
screen "AI" 800x480, template "Main"
   Button "Button_1" at 7,5 size 96x32; TextOff 'Мешалки'; Authorization "Admin"
      on Release: ActivateScreen("Mix", 0); SetTag("settings", 1)
      Appearance <- "settings"
   Button "Button_2" at 7,52 size 96x32; TextOff 'Дозаторы'; Authorization "Admin"
      on Release: ActivateScreen("Dos", 0); SetTag("settings", 2)
      Appearance <- "settings"
   Button "Button_3" at 7,99 size 96x32; TextOff 'Клапана'; Authorization "Admin"
      on Release: ActivateScreen("Valve", 0); SetTag("settings", 3)
      Appearance <- "settings"
   Button "Button_4" at 7,146 size 96x32; TextOff 'AI'; Authorization "Admin"
      on Release: ActivateScreen("AI", 0); SetTag("settings", 4)
      Appearance <- "settings"
   Button "Button_5" at 7,193 size 96x32; TextOff 'DI'; Authorization "Admin"
      on Release: ActivateScreen("DI", 0); SetTag("settings", 5)
      Appearance <- "settings"
   Button "Button_6" at 7,240 size 96x32; TextOff 'DO'; Authorization "Admin"
      on Release: ActivateScreen("DO", 0); SetTag("settings", 6)
      Appearance <- "settings"
   TextField "Text field_2" at 210,15 size 67x22; Text 'Датчик:'
   TextField "Text field_4" at 282,15 size 99x22; Text 'Расходомер'
   TextField "Text field_7" at 390,18 size 43x22; Text 'вход'
   TextField "Text field_8" at 390,43 size 56x22; Text 'выход'
   IOField "I/O field_1" at 456,19 size 92x26; FormatPattern s999999999.999
      ProcessValue <- "AIx_DB_FlowMeter_Converter_Min_In"
   IOField "I/O field_2" at 456,41 size 92x26; FormatPattern s999999999.999
      ProcessValue <- "AIx_DB_FlowMeter_Converter_Min_Out"
   IOField "I/O field_3" at 555,18 size 92x26; FormatPattern s999999999.999
      ProcessValue <- "AIx_DB_FlowMeter_Converter_Max_In"
   IOField "I/O field_4" at 555,40 size 92x26; FormatPattern s999999999.999
      ProcessValue <- "AIx_DB_FlowMeter_Converter_Max_Out"
   TextField "Text field_9" at 389,68 size 101x22; Text 'Фильтрация'
   TextField "Text field_10" at 390,96 size 36x22; Text 'RTD'
   Button "Button_7" at 489,71 size 20x20; TextOff 'Text'; PictureList "ok"
      on Click: InvertBit("AIx_DB_FlowMeter_Use_Filter")
      ProcessValue <- "AIx_DB_FlowMeter_Use_Filter"
   Button "Button_8" at 489,96 size 20x20; TextOff 'Text'; PictureList "ok"
      on Click: InvertBit("AIx_DB_FlowMeter_Use_RTD")
      ProcessValue <- "AIx_DB_FlowMeter_Use_RTD"
   IOField "I/O field_5" at 516,68 size 65x25; FormatPattern 999
      ProcessValue <- "AIx_DB_FlowMeter_Filter_SP"
   IOField "I/O field_6" at 516,93 size 65x25; FormatPattern 999
      ProcessValue <- "AIx_DB_FlowMeter_RTD_c"
   TextField "Text field_11" at 210,36 size 79x22; Text 'Поправка'
   IOField "I/O field_7" at 293,36 size 78x23; FormatPattern s999.9
      ProcessValue <- "AIx_DB_FlowMeter_Calibration"
   Button "Button_9" at 396,176 size 248x28; TextOff 'Use'
      on Click: InvertBit("AIx_DB_FlowMeter_CMD_Start_A")
      Appearance <- "AIx_DB_FlowMeter_CMD_Start_A"
   Button "Button_10" at 213,66 size 68x28; TextOff 'Hand'
      on Click: InvertBit("AIx_DB_FlowMeter_CMD_Hand")
      Appearance <- "AIx_DB_FlowMeter_CMD_Hand"
   IOField "I/O field_8" at 293,66 size 78x28; FormatPattern s9999.9
      ProcessValue <- "AIx_DB_FlowMeter_Result"
   TextField "Text field_12" at 436,123 size 27x22; Text 'NC'
   TextField "Text field_13" at 437,143 size 25x22; Text 'SC'
   TextField "Text field_14" at 210,125 size 27x22; Text 'HH'
   TextField "Text field_15" at 216,145 size 16x22; Text 'H'
   TextField "Text field_16" at 217,165 size 14x22; Text 'L'
   TextField "Text field_17" at 212,186 size 23x22; Text 'LL'
   IOField "I/O field_11" at 472,123 size 58x21; FormatPattern s99999
      ProcessValue <- "AIx_DB_FlowMeter_SP_NC"
   IOField "I/O field_12" at 472,143 size 58x21; FormatPattern s99999
      ProcessValue <- "AIx_DB_FlowMeter_SP_SC"
   IOField "I/O field_13" at 246,125 size 58x21; FormatPattern 99999
      ProcessValue <- "AIx_DB_FlowMeter_SP_HH"
   IOField "I/O field_14" at 246,145 size 58x21; FormatPattern 99999
      ProcessValue <- "AIx_DB_FlowMeter_SP_H"
   IOField "I/O field_15" at 246,165 size 58x21; FormatPattern s99999
      ProcessValue <- "AIx_DB_FlowMeter_SP_L"
   IOField "I/O field_16" at 246,185 size 58x21; FormatPattern s99999
      ProcessValue <- "AIx_DB_FlowMeter_SP_LL"
   IOField "I/O field_17" at 546,123 size 58x21; FormatPattern 999
      ProcessValue <- "AIx_DB_FlowMeter_Timers_NC_SP"
   IOField "I/O field_18" at 546,143 size 58x21; FormatPattern 999
      ProcessValue <- "AIx_DB_FlowMeter_Timers_SC_SP"
   IOField "I/O field_19" at 320,125 size 58x21; FormatPattern 999
      ProcessValue <- "AIx_DB_FlowMeter_Timers_HH_SP"
   IOField "I/O field_20" at 320,145 size 58x21; FormatPattern 999
      ProcessValue <- "AIx_DB_FlowMeter_Timers_H_SP"
   IOField "I/O field_21" at 320,165 size 58x21; FormatPattern 999
      ProcessValue <- "AIx_DB_FlowMeter_Timers_L_SP"
   IOField "I/O field_22" at 320,185 size 58x21; FormatPattern 999
      ProcessValue <- "AIx_DB_FlowMeter_Timers_LL_SP"
   IOField "I/O field_23" at 582,93 size 65x25; FormatPattern s99999
      ProcessValue <- "AIx_DB_FlowMeter_Signal"
   TextField "Text field_18" at 210,97 size 68x22; Text 'Уставка'
   TextField "Text field_19" at 299,97 size 79x22; Text 'Время (с)'
   TextField "Text field_1" at 214,248 size 67x22; Text 'Датчик:'
   TextField "Text field_3" at 286,248 size 69x22; Text 'Уровень'
   TextField "Text field_5" at 394,251 size 43x22; Text 'вход'
   TextField "Text field_6" at 394,276 size 56x22; Text 'выход'
   IOField "I/O field_9" at 460,252 size 92x26; FormatPattern s999999999.999
      ProcessValue <- "AIx_DB_Level_Converter_Min_In"
   IOField "I/O field_10" at 460,274 size 92x26; FormatPattern s999999999.999
      ProcessValue <- "AIx_DB_Level_Converter_Min_Out"
   IOField "I/O field_24" at 559,251 size 92x26; FormatPattern s999999999.999
      ProcessValue <- "AIx_DB_Level_Converter_Max_In"
   IOField "I/O field_25" at 559,273 size 92x26; FormatPattern s999999999.999
      ProcessValue <- "AIx_DB_Level_Converter_Max_Out"
   TextField "Text field_20" at 393,301 size 101x22; Text 'Фильтрация'
   TextField "Text field_21" at 394,329 size 36x22; Text 'RTD'
   Button "Button_11" at 493,304 size 20x20; TextOff 'Text'; PictureList "ok"
      on Click: InvertBit("AIx_DB_Level_Use_Filter")
      ProcessValue <- "AIx_DB_Level_Use_Filter"
   Button "Button_12" at 493,329 size 20x20; TextOff 'Text'; PictureList "ok"
      on Click: InvertBit("AIx_DB_Level_Use_RTD")
      ProcessValue <- "AIx_DB_Level_Use_RTD"
   IOField "I/O field_26" at 520,301 size 65x25; FormatPattern 999
      ProcessValue <- "AIx_DB_Level_Filter_SP"
   IOField "I/O field_27" at 520,326 size 65x25; FormatPattern 999
      ProcessValue <- "AIx_DB_Level_RTD_c"
   TextField "Text field_22" at 214,269 size 79x22; Text 'Поправка'
   IOField "I/O field_28" at 297,269 size 78x23; FormatPattern s999.9
      ProcessValue <- "AIx_DB_Level_Calibration"
   Button "Button_13" at 400,409 size 248x28; TextOff 'Use'
      on Click: InvertBit("AIx_DB_Level_CMD_Start_A")
      Appearance <- "AIx_DB_Level_CMD_Start_A"
   Button "Button_14" at 217,299 size 68x28; TextOff 'Hand'
      on Click: InvertBit("AIx_DB_Level_CMD_Hand")
      Appearance <- "AIx_DB_Level_CMD_Hand"
   IOField "I/O field_29" at 297,299 size 78x28; FormatPattern s9999.9
      ProcessValue <- "AIx_DB_Level_Result"
   TextField "Text field_23" at 440,356 size 27x22; Text 'NC'
   TextField "Text field_24" at 441,376 size 25x22; Text 'SC'
   TextField "Text field_25" at 214,358 size 27x22; Text 'HH'
   TextField "Text field_26" at 220,378 size 16x22; Text 'H'
   TextField "Text field_27" at 221,398 size 14x22; Text 'L'
   TextField "Text field_28" at 216,419 size 23x22; Text 'LL'
   IOField "I/O field_30" at 476,356 size 58x21; FormatPattern s99999
      ProcessValue <- "AIx_DB_Level_SP_NC"
   IOField "I/O field_31" at 476,376 size 58x21; FormatPattern s99999
      ProcessValue <- "AIx_DB_Level_SP_SC"
   IOField "I/O field_32" at 250,358 size 58x21; FormatPattern 99999
      ProcessValue <- "AIx_DB_Level_SP_HH"
   IOField "I/O field_33" at 250,378 size 58x21; FormatPattern 99999
      ProcessValue <- "AIx_DB_Level_SP_H"
   IOField "I/O field_34" at 250,398 size 58x21; FormatPattern s99999
      ProcessValue <- "AIx_DB_Level_SP_L"
   IOField "I/O field_35" at 250,418 size 58x21; FormatPattern s99999
      ProcessValue <- "AIx_DB_Level_SP_LL"
   IOField "I/O field_36" at 550,356 size 58x21; FormatPattern 999
      ProcessValue <- "AIx_DB_Level_Timers_NC_SP"
   IOField "I/O field_37" at 550,376 size 58x21; FormatPattern 999
      ProcessValue <- "AIx_DB_Level_Timers_SC_SP"
   IOField "I/O field_38" at 324,358 size 58x21; FormatPattern 999
      ProcessValue <- "AIx_DB_Level_Timers_HH_SP"
   IOField "I/O field_39" at 324,378 size 58x21; FormatPattern 999
      ProcessValue <- "AIx_DB_Level_Timers_H_SP"
   IOField "I/O field_40" at 324,398 size 58x21; FormatPattern 999
      ProcessValue <- "AIx_DB_Level_Timers_L_SP"
   IOField "I/O field_41" at 324,418 size 58x21; FormatPattern 999
      ProcessValue <- "AIx_DB_Level_Timers_LL_SP"
   IOField "I/O field_42" at 586,326 size 65x25; FormatPattern s99999
      ProcessValue <- "AIx_DB_Level_Signal"
   TextField "Text field_29" at 214,330 size 68x22; Text 'Уставка'
   TextField "Text field_30" at 303,330 size 79x22; Text 'Время (с)'

screen "DI" 800x480, template "Main"
   Button "Button_1" at 7,5 size 96x32; TextOff 'Мешалки'; Authorization "Admin"
      on Release: ActivateScreen("Mix", 0); SetTag("settings", 1)
      Appearance <- "settings"
   Button "Button_2" at 7,52 size 96x32; TextOff 'Дозаторы'; Authorization "Admin"
      on Release: ActivateScreen("Dos", 0); SetTag("settings", 2)
      Appearance <- "settings"
   Button "Button_3" at 7,99 size 96x32; TextOff 'Клапана'; Authorization "Admin"
      on Release: ActivateScreen("Valve", 0); SetTag("settings", 3)
      Appearance <- "settings"
   Button "Button_4" at 7,146 size 96x32; TextOff 'AI'; Authorization "Admin"
      on Release: ActivateScreen("AI", 0); SetTag("settings", 4)
      Appearance <- "settings"
   Button "Button_5" at 7,193 size 96x32; TextOff 'DI'; Authorization "Admin"
      on Release: ActivateScreen("DI", 0); SetTag("settings", 5)
      Appearance <- "settings"
   Button "Button_6" at 7,240 size 96x32; TextOff 'DO'; Authorization "Admin"
      on Release: ActivateScreen("DO", 0); SetTag("settings", 6)
      Appearance <- "settings"
   Group "Group" at 127,7 size 283x51; TextList "Hand"
   Group "Group_1" at 127,66 size 283x51; TextList "Hand"
   Group "Group_2" at 127,125 size 283x51; TextList "Hand"
   Group "Group_3" at 127,184 size 283x51; TextList "Hand"
   Group "Group_4" at 127,244 size 283x51; TextList "Hand"
   Group "Group_5" at 127,303 size 283x51; TextList "Hand"
   Group "Group_6" at 127,362 size 283x51; TextList "Hand"
   Group "Group_7" at 127,422 size 283x51; TextList "Hand"
   Group "Group_8" at 433,7 size 283x51; TextList "Hand"
   Group "Group_9" at 433,66 size 283x51; TextList "Hand"
   Group "Group_10" at 433,125 size 283x51; TextList "Hand"
   Group "Group_11" at 433,184 size 283x51; TextList "Hand"
   Group "Group_12" at 433,244 size 283x51; TextList "Hand"
   Group "Group_13" at 433,303 size 283x51; TextList "Hand"
   TextField "Text field_1" at 131,10 size 45x22; Text 'I 0.0'
   TextField "Text field_2" at 176,10 size 120x22; Text 'M1 Готовность'
   Circle "Circle_1" at 131,33 size 22x22
      Appearance <- "DIx_DB_M1_FB_Ready_Input"
   Circle "Circle_2" at 154,33 size 22x22
      Appearance <- "DIx_DB_M1_FB_Ready_Signal"
   Button "Button_7" at 298,11 size 59x44; TextOff 'Авто'; TextList "Hand"
      on Click: InvertBit("DIx_DB_M1_FB_Ready_Hand")
      Appearance <- "DIx_DB_M1_FB_Ready_Hand"
      ProcessValue <- "DIx_DB_M1_FB_Ready_Hand"
   Button "Button_8" at 240,33 size 49x22; TextOff 'Выкл'
      on Click: ResetBit("DIx_DB_M1_FB_Ready_Start_M")
   Button "Button_12" at 184,33 size 47x22; TextOff 'Вкл'
      on Click: SetBit("DIx_DB_M1_FB_Ready_Start_M")
      Appearance <- "DIx_DB_M1_FB_Ready_Start_M"
   IOField "I/O field_6" at 360,33 size 23x22; FormatPattern 99
      ProcessValue <- "DIx_DB_M1_FB_Ready_Filter_On_SP"
   IOField "I/O field_7" at 383,33 size 23x22; FormatPattern 99
      ProcessValue <- "DIx_DB_M1_FB_Ready_Filter_Off_SP"
   Button "Button_9" at 360,10 size 46x20; TextOff 'Inv'
      on Click: InvertBit("DIx_DB_M1_FB_Ready_Inverse")
      Appearance <- "DIx_DB_M1_FB_Ready_Inverse"
   TextField "Text field_3" at 131,69 size 45x22; Text 'I 0.1'
   TextField "Text field_4" at 176,69 size 87x22; Text 'M1 Работа'
   Circle "Circle_3" at 131,92 size 22x22
      Appearance <- "DIx_DB_M1_FB_Run_Input"
   Circle "Circle_4" at 154,92 size 22x22
      Appearance <- "DIx_DB_M1_FB_Run_Signal"
   Button "Button_10" at 298,70 size 59x44; TextOff 'Авто'; TextList "Hand"
      on Click: InvertBit("DIx_DB_M1_FB_Run_Hand")
      Appearance <- "DIx_DB_M1_FB_Run_Hand"
      ProcessValue <- "DIx_DB_M1_FB_Run_Hand"
   Button "Button_11" at 240,92 size 49x22; TextOff 'Выкл'
      on Click: ResetBit("DIx_DB_M1_FB_Run_Start_M")
   Button "Button_13" at 184,92 size 47x22; TextOff 'Вкл'
      on Click: SetBit("DIx_DB_M1_FB_Run_Start_M")
      Appearance <- "DIx_DB_M1_FB_Run_Start_M"
   IOField "I/O field_1" at 360,92 size 23x22; FormatPattern 99
      ProcessValue <- "DIx_DB_M1_FB_Run_Filter_On_SP"
   IOField "I/O field_2" at 383,92 size 23x22; FormatPattern 99
      ProcessValue <- "DIx_DB_M1_FB_Run_Filter_Off_SP"
   Button "Button_14" at 360,69 size 46x20; TextOff 'Inv'
      on Click: InvertBit("DIx_DB_M1_FB_Run_Inverse")
      Appearance <- "DIx_DB_M1_FB_Run_Inverse"
   TextField "Text field_5" at 131,128 size 45x22; Text 'I 0.2'
   TextField "Text field_6" at 176,128 size 120x22; Text 'M2 Готовность'
   Circle "Circle_5" at 131,151 size 22x22
      Appearance <- "DIx_DB_M2_FB_Ready_Input"
   Circle "Circle_6" at 154,151 size 22x22
      Appearance <- "DIx_DB_M2_FB_Ready_Signal"
   Button "Button_15" at 298,129 size 59x44; TextOff 'Авто'; TextList "Hand"
      on Click: InvertBit("DIx_DB_M2_FB_Ready_Hand")
      Appearance <- "DIx_DB_M2_FB_Ready_Hand"
      ProcessValue <- "DIx_DB_M2_FB_Ready_Hand"
   Button "Button_16" at 240,151 size 49x22; TextOff 'Выкл'
      on Click: ResetBit("DIx_DB_M2_FB_Ready_Start_M")
   Button "Button_17" at 184,151 size 47x22; TextOff 'Вкл'
      on Click: SetBit("DIx_DB_M2_FB_Ready_Start_M")
      Appearance <- "DIx_DB_M2_FB_Ready_Start_M"
   IOField "I/O field_3" at 360,151 size 23x22; FormatPattern 99
      ProcessValue <- "DIx_DB_M2_FB_Ready_Filter_On_SP"
   IOField "I/O field_4" at 383,151 size 23x22; FormatPattern 99
      ProcessValue <- "DIx_DB_M2_FB_Ready_Filter_Off_SP"
   Button "Button_18" at 360,128 size 46x20; TextOff 'Inv'
      on Click: InvertBit("DIx_DB_M2_FB_Ready_Inverse")
      Appearance <- "DIx_DB_M2_FB_Ready_Inverse"
   TextField "Text field_7" at 131,187 size 45x22; Text 'I 0.3'
   TextField "Text field_8" at 176,187 size 87x22; Text 'M2 Работа'
   Circle "Circle_7" at 131,210 size 22x22
      Appearance <- "DIx_DB_M2_FB_Run_Input"
   Circle "Circle_8" at 154,210 size 22x22
      Appearance <- "DIx_DB_M2_FB_Run_Signal"
   Button "Button_19" at 298,188 size 59x44; TextOff 'Авто'; TextList "Hand"
      on Click: InvertBit("DIx_DB_M2_FB_Run_Hand")
      Appearance <- "DIx_DB_M2_FB_Run_Hand"
      ProcessValue <- "DIx_DB_M2_FB_Run_Hand"
   Button "Button_20" at 240,210 size 49x22; TextOff 'Выкл'
      on Click: ResetBit("DIx_DB_M2_FB_Run_Start_M")
   Button "Button_21" at 184,210 size 47x22; TextOff 'Вкл'
      on Click: SetBit("DIx_DB_M2_FB_Run_Start_M")
      Appearance <- "DIx_DB_M2_FB_Run_Start_M"
   IOField "I/O field_5" at 360,210 size 23x22; FormatPattern 99
      ProcessValue <- "DIx_DB_M2_FB_Run_Filter_On_SP"
   IOField "I/O field_8" at 383,210 size 23x22; FormatPattern 99
      ProcessValue <- "DIx_DB_M2_FB_Run_Filter_Off_SP"
   Button "Button_22" at 360,187 size 46x20; TextOff 'Inv'
      on Click: InvertBit("DIx_DB_M2_FB_Run_Inverse")
      Appearance <- "DIx_DB_M2_FB_Run_Inverse"
   TextField "Text field_9" at 131,247 size 45x22; Text 'I 0.4'
   TextField "Text field_10" at 176,247 size 120x22; Text 'M3 Готовность'
   Circle "Circle_9" at 131,270 size 22x22
      Appearance <- "DIx_DB_M3_FB_Ready_Input"
   Circle "Circle_10" at 154,270 size 22x22
      Appearance <- "DIx_DB_M3_FB_Ready_Signal"
   Button "Button_23" at 298,248 size 59x44; TextOff 'Авто'; TextList "Hand"
      on Click: InvertBit("DIx_DB_M3_FB_Ready_Hand")
      Appearance <- "DIx_DB_M3_FB_Ready_Hand"
      ProcessValue <- "DIx_DB_M3_FB_Ready_Hand"
   Button "Button_24" at 240,270 size 49x22; TextOff 'Выкл'
      on Click: ResetBit("DIx_DB_M3_FB_Ready_Start_M")
   Button "Button_25" at 184,270 size 47x22; TextOff 'Вкл'
      on Click: SetBit("DIx_DB_M3_FB_Ready_Start_M")
      Appearance <- "DIx_DB_M3_FB_Ready_Start_M"
   IOField "I/O field_9" at 360,270 size 23x22; FormatPattern 99
      ProcessValue <- "DIx_DB_M3_FB_Ready_Filter_On_SP"
   IOField "I/O field_10" at 383,270 size 23x22; FormatPattern 99
      ProcessValue <- "DIx_DB_M3_FB_Ready_Filter_Off_SP"
   Button "Button_26" at 360,247 size 46x20; TextOff 'Inv'
      on Click: InvertBit("DIx_DB_M3_FB_Ready_Inverse")
      Appearance <- "DIx_DB_M3_FB_Ready_Inverse"
   TextField "Text field_11" at 131,306 size 45x22; Text 'I 0.5'
   TextField "Text field_12" at 176,306 size 87x22; Text 'M3 Работа'
   Circle "Circle_11" at 131,329 size 22x22
      Appearance <- "DIx_DB_M3_FB_Run_Input"
   Circle "Circle_12" at 154,329 size 22x22
      Appearance <- "DIx_DB_M3_FB_Run_Signal"
   Button "Button_27" at 298,307 size 59x44; TextOff 'Авто'; TextList "Hand"
      on Click: InvertBit("DIx_DB_M3_FB_Run_Hand")
      Appearance <- "DIx_DB_M3_FB_Run_Hand"
      ProcessValue <- "DIx_DB_M3_FB_Run_Hand"
   Button "Button_28" at 240,329 size 49x22; TextOff 'Выкл'
      on Click: ResetBit("DIx_DB_M3_FB_Run_Start_M")
   Button "Button_29" at 184,329 size 47x22; TextOff 'Вкл'
      on Click: SetBit("DIx_DB_M3_FB_Run_Start_M")
      Appearance <- "DIx_DB_M3_FB_Run_Start_M"
   IOField "I/O field_11" at 360,329 size 23x22; FormatPattern 99
      ProcessValue <- "DIx_DB_M3_FB_Run_Filter_On_SP"
   IOField "I/O field_12" at 383,329 size 23x22; FormatPattern 99
      ProcessValue <- "DIx_DB_M3_FB_Run_Filter_Off_SP"
   Button "Button_30" at 360,306 size 46x20; TextOff 'Inv'
      on Click: InvertBit("DIx_DB_M3_FB_Run_Inverse")
      Appearance <- "DIx_DB_M3_FB_Run_Inverse"
   TextField "Text field_13" at 131,365 size 45x22; Text 'I 0.6'
   TextField "Text field_14" at 176,365 size 120x22; Text 'Сух.доз.Готов.'
   Circle "Circle_13" at 131,388 size 22x22
      Appearance <- "DIx_DB_DD_FB_Ready_Input"
   Circle "Circle_14" at 154,388 size 22x22
      Appearance <- "DIx_DB_DD_FB_Ready_Signal"
   Button "Button_31" at 298,366 size 59x44; TextOff 'Авто'; TextList "Hand"
      on Click: InvertBit("DIx_DB_DD_FB_Ready_Hand")
      Appearance <- "DIx_DB_DD_FB_Ready_Hand"
      ProcessValue <- "DIx_DB_DD_FB_Ready_Hand"
   Button "Button_32" at 240,388 size 49x22; TextOff 'Выкл'
      on Click: ResetBit("DIx_DB_DD_FB_Ready_Start_M")
   Button "Button_33" at 184,388 size 47x22; TextOff 'Вкл'
      on Click: SetBit("DIx_DB_DD_FB_Ready_Start_M")
      Appearance <- "DIx_DB_DD_FB_Ready_Start_M"
   IOField "I/O field_13" at 360,388 size 23x22; FormatPattern 99
      ProcessValue <- "DIx_DB_DD_FB_Ready_Filter_On_SP"
   IOField "I/O field_14" at 383,388 size 23x22; FormatPattern 99
      ProcessValue <- "DIx_DB_DD_FB_Ready_Filter_Off_SP"
   Button "Button_34" at 360,365 size 46x20; TextOff 'Inv'
      on Click: InvertBit("DIx_DB_DD_FB_Ready_Inverse")
      Appearance <- "DIx_DB_DD_FB_Ready_Inverse"
   TextField "Text field_15" at 131,425 size 45x22; Text 'I 0.7'
   TextField "Text field_16" at 176,425 size 98x22; Text 'Доз. Работа'
   Circle "Circle_15" at 131,448 size 22x22
      Appearance <- "DIx_DB_Dos_FB_Run_Input"
   Circle "Circle_16" at 154,448 size 22x22
      Appearance <- "DIx_DB_Dos_FB_Run_Signal"
   Button "Button_35" at 298,426 size 59x44; TextOff 'Авто'; TextList "Hand"
      on Click: InvertBit("DIx_DB_Dos_FB_Run_Hand")
      ProcessValue <- "DIx_DB_Dos_FB_Run_Hand"
      Appearance <- "DIx_DB_Dos_FB_Run_Hand"
   Button "Button_36" at 240,448 size 49x22; TextOff 'Выкл'
      on Click: ResetBit("DIx_DB_Dos_FB_Run_Start_M")
   Button "Button_37" at 184,448 size 47x22; TextOff 'Вкл'
      on Click: SetBit("DIx_DB_Dos_FB_Run_Start_M")
      Appearance <- "DIx_DB_Dos_FB_Run_Start_M"
   IOField "I/O field_15" at 360,448 size 23x22; FormatPattern 99
      ProcessValue <- "DIx_DB_Dos_FB_Run_Filter_On_SP"
   IOField "I/O field_16" at 383,448 size 23x22; FormatPattern 99
      ProcessValue <- "DIx_DB_Dos_FB_Run_Filter_Off_SP"
   Button "Button_38" at 360,425 size 46x20; TextOff 'Inv'
      on Click: InvertBit("DIx_DB_Dos_FB_Run_Inverse")
      Appearance <- "DIx_DB_Dos_FB_Run_Inverse"
   TextField "Text field_17" at 437,10 size 45x22; Text 'I 1.0'
   TextField "Text field_18" at 482,10 size 95x22; Text 'Сух.доз.Ур.'
   Circle "Circle_17" at 437,33 size 22x22
      Appearance <- "DIx_DB_DD_LLS_Input"
   Circle "Circle_18" at 460,33 size 22x22
      Appearance <- "DIx_DB_DD_LLS_Signal"
   Button "Button_39" at 604,11 size 59x44; TextOff 'Авто'; TextList "Hand"
      on Click: InvertBit("DIx_DB_DD_LLS_Hand")
      Appearance <- "DIx_DB_DD_LLS_Hand"
      ProcessValue <- "DIx_DB_DD_LLS_Hand"
   Button "Button_40" at 546,33 size 49x22; TextOff 'Выкл'
      on Click: ResetBit("DIx_DB_DD_LLS_Start_M")
   Button "Button_41" at 490,33 size 47x22; TextOff 'Вкл'
      on Click: SetBit("DIx_DB_DD_LLS_Start_M")
      Appearance <- "DIx_DB_DD_LLS_Start_M"
   IOField "I/O field_17" at 666,33 size 23x22; FormatPattern 99
      ProcessValue <- "DIx_DB_DD_LLS_Filter_On_SP"
   IOField "I/O field_18" at 689,33 size 23x22; FormatPattern 99
      ProcessValue <- "DIx_DB_DD_LLS_Filter_Off_SP"
   Button "Button_42" at 666,10 size 46x20; TextOff 'Inv'
      on Click: InvertBit("DIx_DB_DD_LLS_Inverse")
      Appearance <- "DIx_DB_DD_LLS_Inverse"
   TextField "Text field_19" at 437,69 size 45x22; Text 'I 1.1'
   TextField "Text field_20" at 482,69 size 104x22; Text 'Вибро Готов.'
   Circle "Circle_19" at 437,92 size 22x22
      Appearance <- "DIx_DB_Vibro_FB_Ready_Input"
   Circle "Circle_20" at 460,92 size 22x22
      Appearance <- "DIx_DB_Vibro_FB_Ready_Signal"
   Button "Button_43" at 604,70 size 59x44; TextOff 'Авто'; TextList "Hand"
      on Click: InvertBit("DIx_DB_Vibro_FB_Ready_Hand")
      Appearance <- "DIx_DB_Vibro_FB_Ready_Hand"
      ProcessValue <- "DIx_DB_Vibro_FB_Ready_Hand"
   Button "Button_44" at 546,92 size 49x22; TextOff 'Выкл'
      on Click: ResetBit("DIx_DB_Vibro_FB_Ready_Start_M")
   Button "Button_45" at 490,92 size 47x22; TextOff 'Вкл'
      on Click: SetBit("DIx_DB_Vibro_FB_Ready_Start_M")
      Appearance <- "DIx_DB_Vibro_FB_Ready_Start_M"
   IOField "I/O field_19" at 666,92 size 23x22; FormatPattern 99
      ProcessValue <- "DIx_DB_Vibro_FB_Ready_Filter_On_SP"
   IOField "I/O field_20" at 689,92 size 23x22; FormatPattern 99
      ProcessValue <- "DIx_DB_Vibro_FB_Ready_Filter_Off_SP"
   Button "Button_46" at 666,69 size 46x20; TextOff 'Inv'
      on Click: InvertBit("DIx_DB_Vibro_FB_Ready_Inverse")
      Appearance <- "DIx_DB_Vibro_FB_Ready_Inverse"
   TextField "Text field_21" at 437,128 size 45x22; Text 'I 1.2'
   TextField "Text field_22" at 482,128 size 112x22; Text 'Пневмотранс.'
   Circle "Circle_21" at 437,151 size 22x22
      Appearance <- "DIx_DB_Transporter_Input"
   Circle "Circle_22" at 460,151 size 22x22
      Appearance <- "DIx_DB_Transporter_Signal"
   Button "Button_47" at 604,129 size 59x44; TextOff 'Авто'; TextList "Hand"
      on Click: InvertBit("DIx_DB_Transporter_Hand")
      Appearance <- "DIx_DB_Transporter_Hand"
      ProcessValue <- "DIx_DB_Transporter_Hand"
   Button "Button_48" at 546,151 size 49x22; TextOff 'Выкл'
      on Click: ResetBit("DIx_DB_Transporter_Start_M")
   Button "Button_49" at 490,151 size 47x22; TextOff 'Вкл'
      on Click: SetBit("DIx_DB_Transporter_Start_M")
      Appearance <- "DIx_DB_Transporter_Start_M"
   IOField "I/O field_21" at 666,151 size 23x22; FormatPattern 99
      ProcessValue <- "DIx_DB_Transporter_Filter_On_SP"
   IOField "I/O field_22" at 689,151 size 23x22; FormatPattern 99
      ProcessValue <- "DIx_DB_Transporter_Filter_Off_SP"
   Button "Button_50" at 666,128 size 46x20; TextOff 'Inv'
      on Click: InvertBit("DIx_DB_Transporter_Inverse")
      Appearance <- "DIx_DB_Transporter_Inverse"
   TextField "Text field_23" at 437,187 size 45x22; Text 'I 1.3'
   TextField "Text field_24" at 482,187 size 128x22; Text 'Жид.доз.Готов.'
   Circle "Circle_23" at 437,210 size 22x22
      Appearance <- "DIx_DB_DL_FB_Ready_Input"
   Circle "Circle_24" at 460,210 size 22x22
      Appearance <- "DIx_DB_DL_FB_Ready_Signal"
   Button "Button_51" at 604,188 size 59x44; TextOff 'Авто'; TextList "Hand"
      on Click: InvertBit("DIx_DB_DL_FB_Ready_Hand")
      Appearance <- "DIx_DB_DL_FB_Ready_Hand"
      ProcessValue <- "DIx_DB_DL_FB_Ready_Hand"
   Button "Button_52" at 546,210 size 49x22; TextOff 'Выкл'
      on Click: ResetBit("DIx_DB_DL_FB_Ready_Start_M")
   Button "Button_53" at 490,210 size 47x22; TextOff 'Вкл'
      on Click: SetBit("DIx_DB_DL_FB_Ready_Start_M")
      Appearance <- "DIx_DB_DL_FB_Ready_Start_M"
   IOField "I/O field_23" at 666,210 size 23x22; FormatPattern 99
      ProcessValue <- "DIx_DB_DL_FB_Ready_Filter_On_SP"
   IOField "I/O field_24" at 689,210 size 23x22; FormatPattern 99
      ProcessValue <- "DIx_DB_DL_FB_Ready_Filter_Off_SP"
   Button "Button_54" at 666,187 size 46x20; TextOff 'Inv'
      on Click: InvertBit("DIx_DB_DL_FB_Ready_Inverse")
      Appearance <- "DIx_DB_DL_FB_Ready_Inverse"
   TextField "Text field_25" at 437,247 size 45x22; Text 'I 1.4'
   TextField "Text field_26" at 482,247 size 61x22; Text 'Проток'
   Circle "Circle_25" at 437,270 size 22x22
      Appearance <- "DIx_DB_Dry_Run_Input"
   Circle "Circle_26" at 460,270 size 22x22
      Appearance <- "DIx_DB_Dry_Run_Signal"
   Button "Button_55" at 604,248 size 59x44; TextOff 'Авто'; TextList "Hand"
      on Click: InvertBit("DIx_DB_Dry_Run_Hand")
      Appearance <- "DIx_DB_Dry_Run_Hand"
      ProcessValue <- "DIx_DB_Dry_Run_Hand"
   Button "Button_56" at 546,270 size 49x22; TextOff 'Выкл'
      on Click: ResetBit("DIx_DB_Dry_Run_Start_M")
   Button "Button_57" at 490,270 size 47x22; TextOff 'Вкл'
      on Click: SetBit("DIx_DB_Dry_Run_Start_M")
      Appearance <- "DIx_DB_Dry_Run_Start_M"
   IOField "I/O field_25" at 666,270 size 23x22; FormatPattern 99
      ProcessValue <- "DIx_DB_Dry_Run_Filter_On_SP"
   IOField "I/O field_26" at 689,270 size 23x22; FormatPattern 99
      ProcessValue <- "DIx_DB_Dry_Run_Filter_Off_SP"
   Button "Button_58" at 666,247 size 46x20; TextOff 'Inv'
      on Click: InvertBit("DIx_DB_Dry_Run_Inverse")
      Appearance <- "DIx_DB_Dry_Run_Inverse"
   TextField "Text field_27" at 437,306 size 45x22; Text 'I 1.5'
   TextField "Text field_28" at 482,306 size 70x22; Text 'Останов'
   Circle "Circle_27" at 437,329 size 22x22
      Appearance <- "DIx_DB_AllBlock_Input"
   Circle "Circle_28" at 460,329 size 22x22
      Appearance <- "DIx_DB_AllBlock_Signal"
   Button "Button_59" at 604,307 size 59x44; TextOff 'Авто'; TextList "Hand"
      on Click: InvertBit("DIx_DB_AllBlock_Hand")
      Appearance <- "DIx_DB_AllBlock_Hand"
      ProcessValue <- "DIx_DB_AllBlock_Hand"
   Button "Button_60" at 546,329 size 49x22; TextOff 'Выкл'
      on Click: ResetBit("DIx_DB_AllBlock_Start_M")
   Button "Button_61" at 490,329 size 47x22; TextOff 'Вкл'
      on Click: SetBit("DIx_DB_AllBlock_Start_M")
      Appearance <- "DIx_DB_AllBlock_Start_M"
   IOField "I/O field_27" at 666,329 size 23x22; FormatPattern 99
      ProcessValue <- "DIx_DB_AllBlock_Filter_On_SP"
   IOField "I/O field_28" at 689,329 size 23x22; FormatPattern 99
      ProcessValue <- "DIx_DB_AllBlock_Filter_Off_SP"
   Button "Button_62" at 666,306 size 46x20; TextOff 'Inv'
      on Click: InvertBit("DIx_DB_AllBlock_Inverse")
      Appearance <- "DIx_DB_AllBlock_Inverse"

screen "DO" 800x480, template "Main"
   Button "Button_1" at 7,5 size 96x32; TextOff 'Мешалки'; Authorization "Admin"
      on Release: ActivateScreen("Mix", 0); SetTag("settings", 1)
      Appearance <- "settings"
   Button "Button_2" at 7,52 size 96x32; TextOff 'Дозаторы'; Authorization "Admin"
      on Release: ActivateScreen("Dos", 0); SetTag("settings", 2)
      Appearance <- "settings"
   Button "Button_3" at 7,99 size 96x32; TextOff 'Клапана'; Authorization "Admin"
      on Release: ActivateScreen("Valve", 0); SetTag("settings", 3)
      Appearance <- "settings"
   Button "Button_4" at 7,146 size 96x32; TextOff 'AI'; Authorization "Admin"
      on Release: ActivateScreen("AI", 0); SetTag("settings", 4)
      Appearance <- "settings"
   Button "Button_5" at 7,193 size 96x32; TextOff 'DI'; Authorization "Admin"
      on Release: ActivateScreen("DI", 0); SetTag("settings", 5)
      Appearance <- "settings"
   Button "Button_6" at 7,240 size 96x32; TextOff 'DO'; Authorization "Admin"
      on Release: ActivateScreen("DO", 0); SetTag("settings", 6)
      Appearance <- "settings"
   Group "Group" at 127,7 size 283x51; TextList "Hand"
   Group "Group_1" at 127,66 size 283x51; Text 'Q 0.0'; TextList "Hand"
   Group "Group_2" at 127,125 size 283x51; Text 'Q 0.0'; TextList "Hand"
   Group "Group_3" at 127,184 size 283x51; Text 'Q 0.0'; TextList "Hand"
   Group "Group_4" at 127,244 size 283x51; Text 'Q 0.0'; TextList "Hand"
   Group "Group_5" at 127,303 size 283x51; Text 'Q 0.0'; TextList "Hand"
   Group "Group_6" at 127,362 size 283x51; Text 'Q 0.0'; TextList "Hand"
   Group "Group_7" at 127,422 size 283x51; Text 'Q 0.0'; TextList "Hand"
   Group "Group_8" at 433,7 size 283x51; Text 'Q 0.0'; TextList "Hand"
   Group "Group_9" at 433,66 size 283x51; Text 'Q 0.0'; TextList "Hand"
   TextField "Text field_4" at 131,10 size 45x22; Text 'Q 0.0'
   TextField "Text field_5" at 176,10 size 69x22; Text 'M1 Пуск'
   Circle "Circle_3" at 131,33 size 22x22
      Appearance <- "DOx_DB_M1_CMD_Start_A"
   Circle "Circle_4" at 154,33 size 22x22
      Appearance <- "DOx_DB_M1_CMD_Q"
   Button "Button_13" at 298,11 size 59x44; TextOff 'Авто'; TextList "Hand"
      on Click: InvertBit("DOx_DB_M1_CMD_Hand")
      Appearance <- "DOx_DB_M1_CMD_Hand"
      ProcessValue <- "DOx_DB_M1_CMD_Hand"
   Button "Button_14" at 240,33 size 49x22; TextOff 'Выкл'
      on Click: ResetBit("DOx_DB_M1_CMD_Start_M")
   Button "Button_15" at 184,33 size 47x22; TextOff 'Вкл'
      on Click: SetBit("DOx_DB_M1_CMD_Start_M")
      Appearance <- "DOx_DB_M1_CMD_Start_M"
   Button "Button_16" at 360,10 size 46x20; TextOff 'Inv'
      on Click: InvertBit("DOx_DB_M1_CMD_Inverse")
      Appearance <- "DOx_DB_M1_CMD_Inverse"
   Button "Button_17" at 360,35 size 46x20; TextOff 'Sim'
      on Click: InvertBit("DOx_DB_M1_CMD_Simulation")
      Appearance <- "DOx_DB_M1_CMD_Simulation"
   TextField "Text field_1" at 131,69 size 45x22; Text 'Q 0.1'
   TextField "Text field_2" at 176,69 size 69x22; Text 'M2 Пуск'
   Circle "Circle_1" at 131,92 size 22x22
      Appearance <- "DOx_DB_M2_CMD_Start_A"
   Circle "Circle_2" at 154,92 size 22x22
      Appearance <- "DOx_DB_M2_CMD_Q"
   Button "Button_7" at 298,70 size 59x44; TextOff 'Авто'; TextList "Hand"
      on Click: InvertBit("DOx_DB_M2_CMD_Hand")
      Appearance <- "DOx_DB_M2_CMD_Hand"
      ProcessValue <- "DOx_DB_M2_CMD_Hand"
   Button "Button_8" at 240,92 size 49x22; TextOff 'Выкл'
      on Click: ResetBit("DOx_DB_M2_CMD_Start_M")
   Button "Button_9" at 184,92 size 47x22; TextOff 'Вкл'
      on Click: SetBit("DOx_DB_M2_CMD_Start_M")
      Appearance <- "DOx_DB_M2_CMD_Start_M"
   Button "Button_10" at 360,69 size 46x20; TextOff 'Inv'
      on Click: InvertBit("DOx_DB_M2_CMD_Inverse")
      Appearance <- "DOx_DB_M2_CMD_Inverse"
   Button "Button_11" at 360,94 size 46x20; TextOff 'Sim'
      on Click: InvertBit("DOx_DB_M2_CMD_Simulation")
      Appearance <- "DOx_DB_M2_CMD_Simulation"
   TextField "Text field_3" at 131,128 size 45x22; Text 'Q 0.2'
   TextField "Text field_6" at 176,128 size 69x22; Text 'M3 Пуск'
   Circle "Circle_5" at 131,151 size 22x22
      Appearance <- "DOx_DB_M3_CMD_Start_A"
   Circle "Circle_6" at 154,151 size 22x22
      Appearance <- "DOx_DB_M3_CMD_Q"
   Button "Button_12" at 298,129 size 59x44; TextOff 'Авто'; TextList "Hand"
      on Click: InvertBit("DOx_DB_M3_CMD_Hand")
      Appearance <- "DOx_DB_M3_CMD_Hand"
      ProcessValue <- "DOx_DB_M3_CMD_Hand"
   Button "Button_18" at 240,151 size 49x22; TextOff 'Выкл'
      on Click: ResetBit("DOx_DB_M3_CMD_Start_M")
   Button "Button_19" at 184,151 size 47x22; TextOff 'Вкл'
      on Click: SetBit("DOx_DB_M3_CMD_Start_M")
      Appearance <- "DOx_DB_M3_CMD_Start_M"
   Button "Button_20" at 360,128 size 46x20; TextOff 'Inv'
      on Click: InvertBit("DOx_DB_M3_CMD_Inverse")
      Appearance <- "DOx_DB_M3_CMD_Inverse"
   Button "Button_21" at 360,153 size 46x20; TextOff 'Sim'
      on Click: InvertBit("DOx_DB_M3_CMD_Simulation")
      Appearance <- "DOx_DB_M3_CMD_Simulation"
   TextField "Text field_7" at 131,187 size 45x22; Text 'Q 0.3'
   TextField "Text field_8" at 176,187 size 109x22; Text 'Сух.Доз.Пуск'
   Circle "Circle_7" at 131,210 size 22x22
      Appearance <- "DOx_DB_DD_CMD_Start_A"
   Circle "Circle_8" at 154,210 size 22x22
      Appearance <- "DOx_DB_DD_CMD_Q"
   Button "Button_22" at 298,188 size 59x44; TextOff 'Авто'; TextList "Hand"
      on Click: InvertBit("DOx_DB_DD_CMD_Hand")
      Appearance <- "DOx_DB_DD_CMD_Hand"
      ProcessValue <- "DOx_DB_DD_CMD_Hand"
   Button "Button_23" at 240,210 size 49x22; TextOff 'Выкл'
      on Click: ResetBit("DOx_DB_DD_CMD_Start_M")
   Button "Button_24" at 184,210 size 47x22; TextOff 'Вкл'
      on Click: SetBit("DOx_DB_DD_CMD_Start_M")
      Appearance <- "DOx_DB_DD_CMD_Start_M"
   Button "Button_25" at 360,187 size 46x20; TextOff 'Inv'
      on Click: InvertBit("DOx_DB_DD_CMD_Inverse")
      Appearance <- "DOx_DB_DD_CMD_Inverse"
   Button "Button_26" at 360,212 size 46x20; TextOff 'Sim'
      on Click: InvertBit("DOx_DB_DD_CMD_Simulation")
      Appearance <- "DOx_DB_DD_CMD_Simulation"
   TextField "Text field_9" at 131,247 size 45x22; Text 'Q 0.4'
   TextField "Text field_10" at 176,247 size 119x22; Text 'Вибратор Пуск'
   Circle "Circle_9" at 131,270 size 22x22
      Appearance <- "DOx_DB_Vibro_CMD_Start_A"
   Circle "Circle_10" at 154,270 size 22x22
      Appearance <- "DOx_DB_Vibro_CMD_Q"
   Button "Button_27" at 298,248 size 59x44; TextOff 'Авто'; TextList "Hand"
      on Click: InvertBit("DOx_DB_Vibro_CMD_Hand")
      Appearance <- "DOx_DB_Vibro_CMD_Hand"
      ProcessValue <- "DOx_DB_Vibro_CMD_Hand"
   Button "Button_28" at 240,270 size 49x22; TextOff 'Выкл'
      on Click: ResetBit("DOx_DB_Vibro_CMD_Start_M")
   Button "Button_29" at 184,270 size 47x22; TextOff 'Вкл'
      on Click: SetBit("DOx_DB_Vibro_CMD_Start_M")
      Appearance <- "DOx_DB_Vibro_CMD_Start_M"
   Button "Button_30" at 360,247 size 46x20; TextOff 'Inv'
      on Click: InvertBit("DOx_DB_Vibro_CMD_Inverse")
      Appearance <- "DOx_DB_Vibro_CMD_Inverse"
   Button "Button_31" at 360,272 size 46x20; TextOff 'Sim'
      on Click: InvertBit("DOx_DB_Vibro_CMD_Simulation")
      Appearance <- "DOx_DB_Vibro_CMD_Simulation"
   TextField "Text field_11" at 131,306 size 45x22; Text 'Q 0.5'
   TextField "Text field_12" at 176,306 size 116x22; Text 'Жид.доз.Пуск'
   Circle "Circle_11" at 131,329 size 22x22
      Appearance <- "DOx_DB_DL_CMD_Start_A"
   Circle "Circle_12" at 154,329 size 22x22
      Appearance <- "DOx_DB_DL_CMD_Q"
   Button "Button_32" at 298,307 size 59x44; TextOff 'Авто'; TextList "Hand"
      on Click: InvertBit("DOx_DB_DL_CMD_Hand")
      Appearance <- "DOx_DB_DL_CMD_Hand"
      ProcessValue <- "DOx_DB_DL_CMD_Hand"
   Button "Button_33" at 240,329 size 49x22; TextOff 'Выкл'
      on Click: ResetBit("DOx_DB_DL_CMD_Start_M")
   Button "Button_34" at 184,329 size 47x22; TextOff 'Вкл'
      on Click: SetBit("DOx_DB_DL_CMD_Start_M")
      Appearance <- "DOx_DB_DL_CMD_Start_M"
   Button "Button_35" at 360,306 size 46x20; TextOff 'Inv'
      on Click: InvertBit("DOx_DB_DL_CMD_Inverse")
      Appearance <- "DOx_DB_DL_CMD_Inverse"
   Button "Button_36" at 360,331 size 46x20; TextOff 'Sim'
      on Click: InvertBit("DOx_DB_DL_CMD_Simulation")
      Appearance <- "DOx_DB_DL_CMD_Simulation"
   TextField "Text field_13" at 131,365 size 45x22; Text 'Q 0.6'
   TextField "Text field_14" at 176,365 size 110x22; Text 'КС1 Открыть'
   Circle "Circle_13" at 131,388 size 22x22
      Appearance <- "DOx_DB_KC1_CMD_Start_A"
   Circle "Circle_14" at 154,388 size 22x22
      Appearance <- "DOx_DB_KC1_CMD_Q"
   Button "Button_37" at 298,366 size 59x44; TextOff 'Авто'; TextList "Hand"
      on Click: InvertBit("DOx_DB_KC1_CMD_Hand")
      Appearance <- "DOx_DB_KC1_CMD_Hand"
      ProcessValue <- "DOx_DB_KC1_CMD_Hand"
   Button "Button_38" at 240,388 size 49x22; TextOff 'Выкл'
      on Click: ResetBit("DOx_DB_KC1_CMD_Start_M")
   Button "Button_39" at 184,388 size 47x22; TextOff 'Вкл'
      on Click: SetBit("DOx_DB_KC1_CMD_Start_M")
      Appearance <- "DOx_DB_KC1_CMD_Start_M"
   Button "Button_40" at 360,365 size 46x20; TextOff 'Inv'
      on Click: InvertBit("DOx_DB_KC1_CMD_Inverse")
      Appearance <- "DOx_DB_KC1_CMD_Inverse"
   Button "Button_41" at 360,390 size 46x20; TextOff 'Sim'
      on Click: InvertBit("DOx_DB_KC1_CMD_Simulation")
      Appearance <- "DOx_DB_KC1_CMD_Simulation"
   TextField "Text field_15" at 131,425 size 45x22; Text 'Q 0.7'
   TextField "Text field_16" at 176,425 size 117x22; Text 'LED Сухой ход'
   Circle "Circle_15" at 131,448 size 22x22
      Appearance <- "DOx_DB_LED_Dry_Run_Start_A"
   Circle "Circle_16" at 154,448 size 22x22
      Appearance <- "DOx_DB_LED_Dry_Run_Q"
   Button "Button_42" at 298,426 size 59x44; TextOff 'Авто'; TextList "Hand"
      on Click: InvertBit("DOx_DB_LED_Dry_Run_Hand")
      Appearance <- "DOx_DB_LED_Dry_Run_Hand"
      ProcessValue <- "DOx_DB_LED_Dry_Run_Hand"
   Button "Button_43" at 240,448 size 49x22; TextOff 'Выкл'
      on Click: ResetBit("DOx_DB_LED_Dry_Run_Start_M")
   Button "Button_44" at 184,448 size 47x22; TextOff 'Вкл'
      on Click: SetBit("DOx_DB_LED_Dry_Run_Start_M")
      Appearance <- "DOx_DB_LED_Dry_Run_Start_M"
   Button "Button_45" at 360,425 size 46x20; TextOff 'Inv'
      on Click: InvertBit("DOx_DB_LED_Dry_Run_Inverse")
      Appearance <- "DOx_DB_LED_Dry_Run_Inverse"
   Button "Button_46" at 360,450 size 46x20; TextOff 'Sim'
      on Click: InvertBit("DOx_DB_LED_Dry_Run_Simulation")
      Appearance <- "DOx_DB_LED_Dry_Run_Simulation"
   TextField "Text field_17" at 437,10 size 45x22; Text 'Q 1.0'
   TextField "Text field_18" at 482,10 size 93x22; Text 'LED Авария'
   Circle "Circle_17" at 437,33 size 22x22
      Appearance <- "DOx_DB_LED_Alarm_Start_A"
   Circle "Circle_18" at 460,33 size 22x22
      Appearance <- "DOx_DB_LED_Alarm_Q"
   Button "Button_47" at 604,11 size 59x44; TextOff 'Авто'; TextList "Hand"
      on Click: InvertBit("DOx_DB_LED_Alarm_Hand")
      Appearance <- "DOx_DB_LED_Alarm_Hand"
      ProcessValue <- "DOx_DB_LED_Alarm_Hand"
   Button "Button_48" at 546,33 size 49x22; TextOff 'Выкл'
      on Click: ResetBit("DOx_DB_LED_Alarm_Start_M")
   Button "Button_49" at 490,33 size 47x22; TextOff 'Вкл'
      on Click: SetBit("DOx_DB_LED_Alarm_Start_M")
      Appearance <- "DOx_DB_LED_Alarm_Start_M"
   Button "Button_50" at 666,10 size 46x20; TextOff 'Inv'
      on Click: InvertBit("DOx_DB_LED_Alarm_Inverse")
      Appearance <- "DOx_DB_LED_Alarm_Inverse"
   Button "Button_51" at 666,35 size 46x20; TextOff 'Sim'
      on Click: InvertBit("DOx_DB_LED_Alarm_Simulation")
      Appearance <- "DOx_DB_LED_Alarm_Simulation"
   TextField "Text field_19" at 437,69 size 45x22; Text 'Q 1.1'
   TextField "Text field_20" at 482,69 size 84x22; Text 'LED Пусто'
   Circle "Circle_19" at 437,92 size 22x22
      Appearance <- "DOx_DB_LED_Empty_Start_A"
   Circle "Circle_20" at 460,92 size 22x22
      Appearance <- "DOx_DB_LED_Empty_Q"
   Button "Button_52" at 604,70 size 59x44; TextOff 'Авто'; TextList "Hand"
      on Click: InvertBit("DOx_DB_LED_Empty_Hand")
      Appearance <- "DOx_DB_LED_Empty_Hand"
      ProcessValue <- "DOx_DB_LED_Empty_Hand"
   Button "Button_53" at 546,92 size 49x22; TextOff 'Выкл'
      on Click: ResetBit("DOx_DB_LED_Empty_Start_M")
   Button "Button_54" at 490,92 size 47x22; TextOff 'Вкл'
      on Click: SetBit("DOx_DB_LED_Empty_Start_M")
      Appearance <- "DOx_DB_LED_Empty_Start_M"
   Button "Button_55" at 666,69 size 46x20; TextOff 'Inv'
      on Click: InvertBit("DOx_DB_LED_Empty_Inverse")
      Appearance <- "DOx_DB_LED_Empty_Inverse"
   Button "Button_56" at 666,94 size 46x20; TextOff 'Sim'
      on Click: InvertBit("DOx_DB_LED_Empty_Simulation")
      Appearance <- "DOx_DB_LED_Empty_Simulation"

screen "About" 800x480, template "Main"
   TextField "Text field_1" at 174,5 size 426x47; Text 'ООО "Водообработка"'
   TextField "Text field_4" at 61,89 size 652x73; Text 'Разработка и поставка оборудования для подготовки реагентов, дозирования, ввода и высокоэффективного перемешивания веществ в непрерывных технологическихх процессах.'
   TextField "Text field_2" at 43,199 size 689x50; Text 'Контактная информация: Адрес: Россия, г. Москва, 111116 ул. Лефортовский вал, д. 7Г, стр. 5'
   TextField "Text field_3" at 238,286 size 299x27; Text 'Телефон: +7 (495) 763-29-73'
   TextField "Text field_5" at 235,313 size 301x27; Text 'http://www.vodoobrabotka.ru'
   GraphicView "Graphic view_1" at 240,358 size 302x96; Picture "logo"

screen "Configuration" 800x480, template "Main"
   GraphicView "Graphic view_2" at 20,174 size 347x286; Picture "clean2"
   GraphicView "Graphic view_1" at 20,61 size 347x209; Picture "clean2"
   TextField "Text field_2" at 97,75 size 192x33; Text 'Конфигурация'
   TextField "Text field_15" at 33,148 size 146x23; Text 'Жидкий дозатор'
   Button "Button_2" at 224,197 size 100x30; TextOff 'Text'; Authorization "Admin"; PictureList "ON_OFF"
      on Click: InvertBit("CONFIG_Config_Use_DD"); ResetBit("CONFIG_Config_Use_DL")
      ProcessValue <- "CONFIG_Config_Use_DD"
   TextField "Text field_1" at 235,5 size 337x47; Text 'Состав установки'
   TextField "Text field_3" at 33,200 size 128x23; Text 'Сухой дозатор'
   Button "Button_1" at 224,145 size 100x30; TextOff 'Text'; Authorization "Admin"; PictureList "ON_OFF"
      on Click: InvertBit("CONFIG_Config_Use_DL"); ResetBit("CONFIG_Config_Use_DD")
      ProcessValue <- "CONFIG_Config_Use_DL"
   TextField "Text field_4" at 48,282 size 99x23; Text 'Мешалка 1'
   Button "Button_3" at 224,331 size 100x30; TextOff 'Text'; Authorization "Admin"; PictureList "ON_OFF"
      on Click: InvertBit("CONFIG_Config_Use_Mix_2")
      ProcessValue <- "CONFIG_Config_Use_Mix_2"
   TextField "Text field_5" at 48,334 size 99x23; Text 'Мешалка 2'
   Button "Button_4" at 224,279 size 100x30; TextOff 'Text'; Authorization "Admin"; PictureList "ON_OFF"
      on Click: InvertBit("CONFIG_Config_Use_Mix_1")
      ProcessValue <- "CONFIG_Config_Use_Mix_1"
   Button "Button_5" at 224,387 size 100x30; TextOff 'Text'; Authorization "Admin"; PictureList "ON_OFF"
      on Click: InvertBit("CONFIG_Config_Use_Mix_3")
      ProcessValue <- "CONFIG_Config_Use_Mix_3"
   TextField "Text field_6" at 48,390 size 99x23; Text 'Мешалка 3'

screen "Settings" 800x480, template "Main"
   Button "Button_1" at 7,5 size 96x32; TextOff 'Мешалки'; Authorization "Admin"
      on Release: ActivateScreen("Mix", 0); SetTag("settings", 1)
      Appearance <- "settings"
   Button "Button_2" at 7,52 size 96x32; TextOff 'Дозаторы'; Authorization "Admin"
      on Release: ActivateScreen("Dos", 0); SetTag("settings", 2)
      Appearance <- "settings"
   Button "Button_3" at 7,99 size 96x32; TextOff 'Клапана'; Authorization "Admin"
      on Release: ActivateScreen("Valve", 0); SetTag("settings", 3)
      Appearance <- "settings"
   Button "Button_4" at 7,146 size 96x32; TextOff 'AI'; Authorization "Admin"
      on Release: ActivateScreen("AI", 0); SetTag("settings", 4)
      Appearance <- "settings"
   Button "Button_5" at 7,193 size 96x32; TextOff 'DI'; Authorization "Admin"
      on Release: ActivateScreen("DI", 0); SetTag("settings", 5)
      Appearance <- "settings"
   Button "Button_6" at 7,240 size 96x32; TextOff 'DO'; Authorization "Admin"
      on Release: ActivateScreen("DO", 0); SetTag("settings", 6)
      Appearance <- "settings"

Template "Main" 800x480
   Button "Button_1" at 735,5 size 60x60; TextOff 'Text'; PictureOff "home_2"
      on Click: ActivateScreen("Root screen", 0)
   Button "Button_2" at 735,72 size 60x60; TextOff 'Text'; PictureOff "sett"
      on Click: ActivateScreen("SP", 0)
   Button "Button_3" at 735,140 size 60x60; TextOff 'Text'; PictureOff "dos_1"
      on Click: ActivateScreen("Calibration", 0)
   Button "Button_4" at 735,207 size 60x60; TextOff 'Text'; PictureOff "sett_1"
      on Click: ActivateScreen("Monitor", 0)
   Button "Button_5" at 735,275 size 60x60; TextOff 'Text'; PictureOff "home_1"; PictureList "Alarm"
      on Click: ActivateScreen("Alarms", 0)
      ProcessValue <- "Any_Alm"
   Button "Button_6" at 735,342 size 60x60; TextOff 'Text'; PictureOff "back"
      on Click: function_efd93a16()
   Button "Button_7" at 735,410 size 60x60; TextOff 'Text'; PictureOff "reset"
      on Click: SetBit("Reset_All")
*)

(* ===== HMI "HMI_RT_3" =====
system functions are stored by id; their names below are inferred from use
connection "HMI_Connection_4": ETHERNET, SMART_S7_1200_OMS

HMI tags "Default tag table"
   "Comm_1_DB_Mix_3_Status" : Int = PLC Comm_1_DB.Mix_3_Status AT %DB11.DBW24, 1 s
   "Comm_1_DB_Mix_2_Status" : Int = PLC Comm_1_DB.Mix_2_Status AT %DB11.DBW18, 1 s
   "Comm_1_DB_Mix_1_Status" : Int = PLC Comm_1_DB.Mix_1_Status AT %DB11.DBW12, 1 s
   "Comm_1_DB_Level" : Real = PLC Comm_1_DB.Level AT %DB11.DBD38, 1 s
   "Comm_2_DB_Level" : Real = PLC Comm_2_DB.Level AT %DB12.DBD38, 1 s
   "Comm_2_DB_Mix_1_Status" : Int = PLC Comm_2_DB.Mix_1_Status AT %DB12.DBW12, 1 s
   "Comm_2_DB_Mix_2_Status" : Int = PLC Comm_2_DB.Mix_2_Status AT %DB12.DBW18, 1 s
   "Comm_2_DB_Mix_3_Status" : Int = PLC Comm_2_DB.Mix_3_Status AT %DB12.DBW24, 1 s
   "Any_Hand" : Bool = PLC Any_Hand AT %M5.0, 1 s
   "Logick_DB_Start" : Bool = PLC Logick_DB.Start AT %DB1.DBX0.0, 1 s
   "Logick_DB_Hand" : Bool = PLC Logick_DB.Hand AT %DB1.DBX0.1, 1 s
   "Logick_DB_Use_M1" : Bool = PLC Logick_DB.Use_M1 AT %DB1.DBX0.6, 1 s
   "Logick_DB_Use_M3" : Bool = PLC Logick_DB.Use_M3 AT %DB1.DBX1.0, 1 s
   "Logick_DB_REQ_M2_1" : Bool = PLC Logick_DB.REQ_M2_1 AT %DB1.DBX1.3, 1 s
   "Logick_DB_Res_M1" : Bool = PLC Logick_DB.Res_M1 AT %DB1.DBX1.1, 1 s
   "Logick_DB_Res_M3" : Bool = PLC Logick_DB.Res_M3 AT %DB1.DBX1.2, 1 s
   "RS232_DB_Mass_1" : Real = PLC RS232_DB.Mass_1 AT %DB2.DBD0, 1 s
   "Statistics_DB_Today_1" : Real = PLC Statistics_DB.Today_1 AT %DB4.DBD40, 1 s
   "Statistics_DB_Mass_2" : Real = PLC Statistics_DB.Mass_2 AT %DB4.DBD4, 1 s
   "Statistics_DB_Mass_1" : Real = PLC Statistics_DB.Mass_1 AT %DB4.DBD0, 1 s
   "Statistics_DB_Today_2" : Real = PLC Statistics_DB.Today_2 AT %DB4.DBD44, 1 s
   "Logick_DB_Fix_1" : Bool = PLC Logick_DB.Fix_1 AT %DB1.DBX0.2, 1 s
   "Logick_DB_Fix_D_1" : Real = PLC Logick_DB.Fix_D_1 AT %DB1.DBD48, 1 s
   "Logick_DB_D_1" : Real = PLC Logick_DB.D_1 AT %DB1.DBD56, 1 s
   "Logick_DB_Fix_2" : Bool = PLC Logick_DB.Fix_2 AT %DB1.DBX0.3, 1 s
   "Logick_DB_Fix_D_2" : Real = PLC Logick_DB.Fix_D_2 AT %DB1.DBD52, 1 s
   "Logick_DB_D_2" : Real = PLC Logick_DB.D_2 AT %DB1.DBD60, 1 s
   "Comm_1_DB_Warning" : Bool = PLC Comm_1_DB.Warning AT %DB11.DBX48.2, 1 s
   "Comm_2_DB_Warning" : Bool = PLC Comm_2_DB.Warning AT %DB12.DBX48.2, 1 s
   "Logick_DB_C_1" : Real = PLC Logick_DB.C_1 AT %DB1.DBD64, 1 s
   "Logick_DB_C_2" : Real = PLC Logick_DB.C_2 AT %DB1.DBD68, 1 s
   "Statistics_DB_Zero_1" : Real = PLC Statistics_DB.Zero_1 AT %DB4.DBD64, 1 s
   "RS232_DB_Mass_2" : Real = PLC RS232_DB.Mass_2 AT %DB2.DBD4, 1 s
   "Statistics_DB_Zero_2" : Real = PLC Statistics_DB.Zero_2 AT %DB4.DBD68, 1 s
   "Statistics_DB_Last_1" : Real = PLC Statistics_DB.Last_1 AT %DB4.DBD24, 1 s
   "Statistics_DB_Delta_1" : Real = PLC Statistics_DB.Delta_1 AT %DB4.DBD32, 1 s
   "Statistics_DB_Max_D_1" : Real = PLC Statistics_DB.Max_D_1 AT %DB4.DBD16, 1 s
   "Statistics_DB_Min_D_1" : Real = PLC Statistics_DB.Min_D_1 AT %DB4.DBD8, 1 s
   "Statistics_DB_T_SP_M" : Int = PLC Statistics_DB.T.SP_M AT %DB4.DBW580, 1 s
   "Statistics_DB_T_SP_S" : Int = PLC Statistics_DB.T.SP_S AT %DB4.DBW582, 1 s
   "Sync" : Bool = PLC Sync_1 AT %M10.0, 1 s
   "Sync_2" : Bool = PLC Sync_2 AT %M10.1, 1 s
   "Statistics_DB_Delta_2" : Real = PLC Statistics_DB.Delta_2 AT %DB4.DBD36, 1 s
   "Statistics_DB_Last_2" : Real = PLC Statistics_DB.Last_2 AT %DB4.DBD28, 1 s
   "Statistics_DB_Max_D_2" : Real = PLC Statistics_DB.Max_D_2 AT %DB4.DBD20, 1 s
   "Statistics_DB_Min_D_2" : Real = PLC Statistics_DB.Min_D_2 AT %DB4.DBD12, 1 s
   "DIx_DB_Heat_4_Signal" : Bool = PLC DIx_DB.Heat_4.Signal AT %DB200.DBX122.0, 1 s
   "DIx_DB_Heat_4_Input" : Bool = PLC DIx_DB.Heat_4.Input AT %DB200.DBX120.0, 1 s
   "DIx_DB_Heat_1_Inverse" : Bool = PLC DIx_DB.Heat_1.Inverse AT %DB200.DBX64.3, 1 s
   "Any_Alm" : Bool = PLC Any_Alm AT %M6.0, 1 s
   "Statistics_DB_Today_Int" : Int = PLC Statistics_DB.Today_Int AT %DB4.DBW74, 1 s
   "Time_Save" : Bool = PLC "Time".Save AT %DB13.DBX38.0, 1 s
   "Time_Year" : UInt = PLC "Time".Year AT %DB13.DBW28, 1 s
   "Time_Month" : UInt = PLC "Time".Month AT %DB13.DBW30, 1 s
   "Time_Day" : UInt = PLC "Time".Day AT %DB13.DBW32, 1 s
   "Time_Hour" : UInt = PLC "Time".Hour AT %DB13.DBW34, 1 s
   "Time_Minutes" : UInt = PLC "Time".Minutes AT %DB13.DBW36, 1 s
   "Time_Today_YEAR" : UInt = PLC "Time".Today.YEAR AT %DB13.DBW0, 1 s
   "Time_Today_MONTH" : USInt = PLC "Time".Today.MONTH AT %DB13.DBB2, 1 s
   "Time_Today_DAY" : USInt = PLC "Time".Today.DAY AT %DB13.DBB3, 1 s
   "Time_Today_WEEKDAY" : USInt = PLC "Time".Today.WEEKDAY AT %DB13.DBB4, 1 s
   "Time_Today_HOUR" : USInt = PLC "Time".Today.HOUR AT %DB13.DBB5, 1 s
   "Time_Today_MINUTE" : USInt = PLC "Time".Today.MINUTE AT %DB13.DBB6, 1 s
   "Reset_All" : Bool = PLC Reset_All AT %M3.1, 1 s
   "Logick_DB_Low_REQ" : Bool = PLC Logick_DB.Low_REQ AT %DB1.DBX2.0, 1 s
   "Logick_DB_Low_view" : Bool = PLC Logick_DB.Low_view AT %DB1.DBX2.2, 1 s
   "Logick_DB_Low_SP_M" : Int = PLC Logick_DB.Low.SP_M AT %DB1.DBW72, 1 s
   "Logick_DB_Low_CMD" : Bool = PLC Logick_DB.Low_CMD AT %DB1.DBX2.1, 1 s
   "Logick_DB_Max_SP" : Real = PLC Logick_DB.Max_SP AT %DB1.DBD36, 1 s
   "Logick_DB_Min_SP" : Real = PLC Logick_DB.Min_SP AT %DB1.DBD32, 1 s
   "Logick_DB_Low_use" : Bool = PLC Logick_DB.Low_use AT %DB1.DBX1.7, 1 s
   "Logick_DB_Correction_1" : Bool = PLC Logick_DB.Correction_1 AT %DB1.DBX2.3, 1 s
   "Logick_DB_Correction_2" : Bool = PLC Logick_DB.Correction_2 AT %DB1.DBX2.4, 1 s
   "Logick_DB_C_SP_1" : Real = PLC Logick_DB.C_SP_1 AT %DB1.DBD40, 1 s
   "Logick_DB_C_SP_2" : Real = PLC Logick_DB.C_SP_2 AT %DB1.DBD44, 1 s

HMI tags "HMI"
   "settings" : Int, internal

